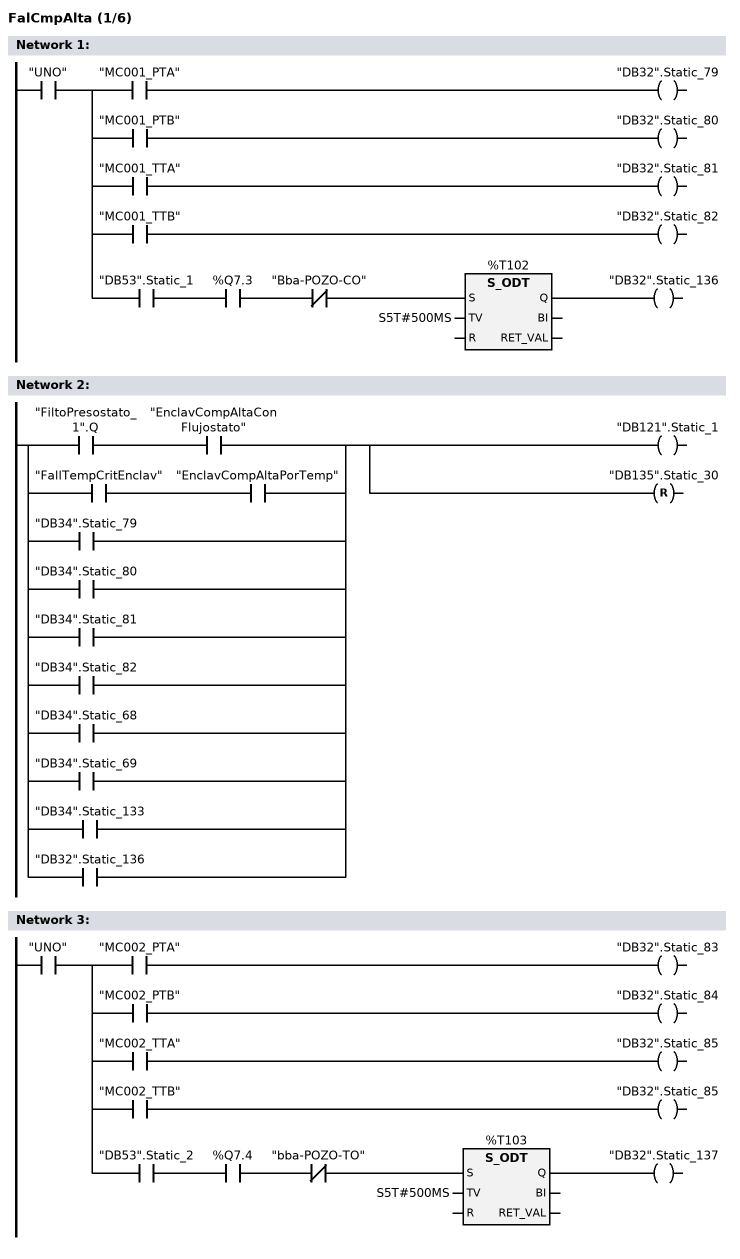
   RUNG wire#powerrail
      Contact( "UNO" )
      wire#w1
      Contact( "MC001_PTA" )
      Coil( "DB32".Static_79 )
   END_RUNG
   RUNG wire#w1
      Contact( "MC001_PTB" )
      Coil( "DB32".Static_80 )
   END_RUNG
   RUNG wire#w1
      Contact( "MC001_TTA" )
      Coil( "DB32".Static_81 )
   END_RUNG
   RUNG wire#w1
      Contact( "MC001_TTB" )
      Coil( "DB32".Static_82 )
   END_RUNG
   RUNG wire#w1
      Contact( "DB53".Static_1 )
      Contact( %Q7.3 )
      I_Contact( "Bba-POZO-CO" )
      S_ODT(T_NO := %T102, TV := S5T#500MS, R :=, BI =>, RET_VAL =>)
      Coil( "DB32".Static_136 )
   END_RUNG
   // the same network as SCL:
   "DB32".Static_79 := "UNO" AND "MC001_PTA";
   "DB32".Static_80 := "UNO" AND "MC001_PTB";
   "DB32".Static_81 := "UNO" AND "MC001_TTA";
   "DB32".Static_82 := "UNO" AND "MC001_TTB";
   #_s5time1 := S_ODT(T_NO := %T102,
                      TV := S5T#500MS,
                      S := "UNO" AND "DB53".Static_1 AND %Q7.3 AND NOT "Bba-POZO-CO",
                      Q => #_w1);
   "DB32".Static_136 := #_w1;
END_REGION

REGION Network 2
   "DB121".Static_1 := "DB34".Static_79 OR "DB34".Static_80 OR "DB34".Static_81 OR "DB34".Static_82 OR "DB34".Static_68 OR "DB34".Static_69 OR "DB34".Static_133 OR ("FiltoPresostato_1".Q AND "EnclavCompAltaConFlujostato") OR ("FallTempCritEnclav" AND "EnclavCompAltaPorTemp") OR "DB32".Static_136;
   IF "DB121".Static_1 THEN "DB135".Static_30 := FALSE; END_IF;
END_REGION

REGION Network 3
   RUNG wire#powerrail
      Contact( "UNO" )
      wire#w1
      Contact( "MC002_PTA" )
      Coil( "DB32".Static_83 )
   END_RUNG
   RUNG wire#w1
      Contact( "MC002_PTB" )
      Coil( "DB32".Static_84 )
   END_RUNG
   RUNG wire#w1
      Contact( "MC002_TTA" )
      Coil( "DB32".Static_85 )
   END_RUNG
   RUNG wire#w1
      Contact( "MC002_TTB" )
      Coil( "DB32".Static_85 )
   END_RUNG
   RUNG wire#w1
      Contact( "DB53".Static_2 )
      Contact( %Q7.4 )
      I_Contact( "bba-POZO-TO" )
      S_ODT(T_NO := %T103, TV := S5T#500MS, R :=, BI =>, RET_VAL =>)
      Coil( "DB32".Static_137 )
   END_RUNG
   // the same network as SCL:
   "DB32".Static_83 := "UNO" AND "MC002_PTA";
   "DB32".Static_84 := "UNO" AND "MC002_PTB";
   "DB32".Static_85 := "UNO" AND "MC002_TTA";
   "DB32".Static_85 := "UNO" AND "MC002_TTB";
   #_s5time1 := S_ODT(T_NO := %T103,
                      TV := S5T#500MS,
                      S := "UNO" AND "DB53".Static_2 AND %Q7.4 AND NOT "bba-POZO-TO",
                      Q => #_w1);
   "DB32".Static_137 := #_w1;
END_REGION

REGION Network 4
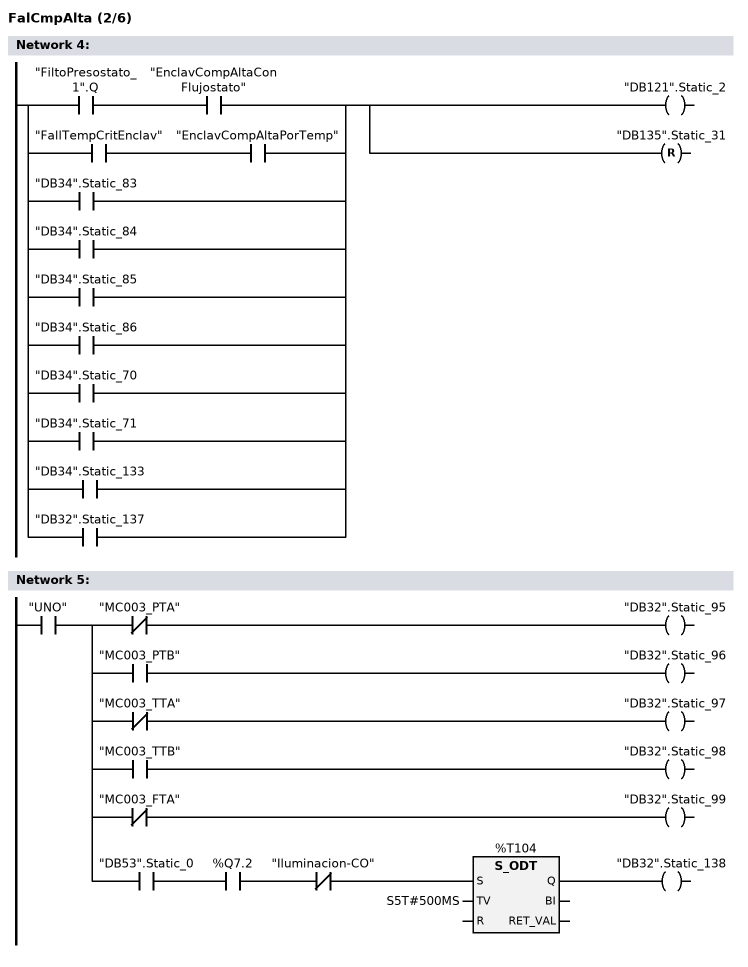
   "DB121".Static_2 := "DB34".Static_83 OR "DB34".Static_84 OR "DB34".Static_85 OR "DB34".Static_86 OR "DB34".Static_70 OR "DB34".Static_71 OR "DB34".Static_133 OR ("FiltoPresostato_1".Q AND "EnclavCompAltaConFlujostato") OR ("FallTempCritEnclav" AND "EnclavCompAltaPorTemp") OR "DB32".Static_137;
   IF "DB121".Static_2 THEN "DB135".Static_31 := FALSE; END_IF;
END_REGION

REGION Network 5
   RUNG wire#powerrail
      Contact( "UNO" )
      wire#w1
      I_Contact( "MC003_PTA" )
      Coil( "DB32".Static_95 )
   END_RUNG
   RUNG wire#w1
      Contact( "MC003_PTB" )
      Coil( "DB32".Static_96 )
   END_RUNG
   RUNG wire#w1
      I_Contact( "MC003_TTA" )
      Coil( "DB32".Static_97 )
   END_RUNG
   RUNG wire#w1
      Contact( "MC003_TTB" )
      Coil( "DB32".Static_98 )
   END_RUNG
   RUNG wire#w1
      I_Contact( "MC003_FTA" )
      Coil( "DB32".Static_99 )
   END_RUNG
   RUNG wire#w1
      Contact( "DB53".Static_0 )
      Contact( %Q7.2 )
      I_Contact( "Iluminacion-CO" )
      S_ODT(T_NO := %T104, TV := S5T#500MS, R :=, BI =>, RET_VAL =>)
      Coil( "DB32".Static_138 )
   END_RUNG
   // the same network as SCL:
   "DB32".Static_95 := "UNO" AND NOT "MC003_PTA";
   "DB32".Static_96 := "UNO" AND "MC003_PTB";
   "DB32".Static_97 := "UNO" AND NOT "MC003_TTA";
   "DB32".Static_98 := "UNO" AND "MC003_TTB";
   "DB32".Static_99 := "UNO" AND NOT "MC003_FTA";
   #_s5time1 := S_ODT(T_NO := %T104,
                      TV := S5T#500MS,
                      S := "UNO" AND "DB53".Static_0 AND %Q7.2 AND NOT "Iluminacion-CO",
                      Q => #_w1);
   "DB32".Static_138 := #_w1;
END_REGION

REGION Network 6
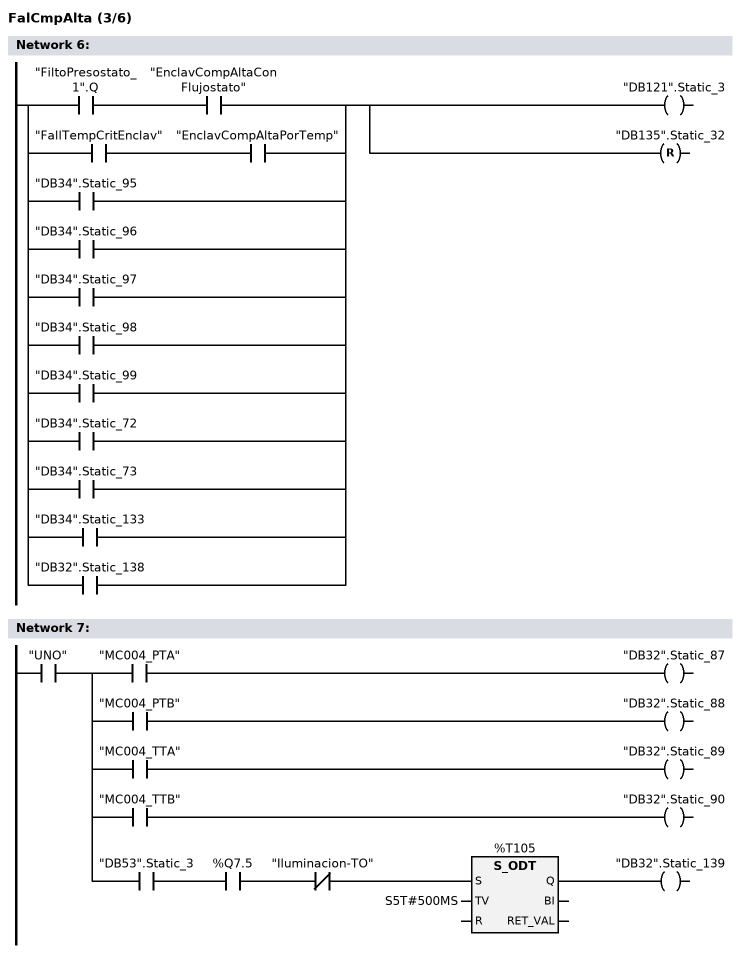
   "DB121".Static_3 := "DB34".Static_95 OR "DB34".Static_96 OR "DB34".Static_97 OR "DB34".Static_98 OR "DB34".Static_99 OR "DB34".Static_72 OR "DB34".Static_73 OR "DB34".Static_133 OR ("FiltoPresostato_1".Q AND "EnclavCompAltaConFlujostato") OR ("FallTempCritEnclav" AND "EnclavCompAltaPorTemp") OR "DB32".Static_138;
   IF "DB121".Static_3 THEN "DB135".Static_32 := FALSE; END_IF;
END_REGION

REGION Network 7
   RUNG wire#powerrail
      Contact( "UNO" )
      wire#w1
      Contact( "MC004_PTA" )
      Coil( "DB32".Static_87 )
   END_RUNG
   RUNG wire#w1
      Contact( "MC004_PTB" )
      Coil( "DB32".Static_88 )
   END_RUNG
   RUNG wire#w1
      Contact( "MC004_TTA" )
      Coil( "DB32".Static_89 )
   END_RUNG
   RUNG wire#w1
      Contact( "MC004_TTB" )
      Coil( "DB32".Static_90 )
   END_RUNG
   RUNG wire#w1
      Contact( "DB53".Static_3 )
      Contact( %Q7.5 )
      I_Contact( "Iluminacion-TO" )
      S_ODT(T_NO := %T105, TV := S5T#500MS, R :=, BI =>, RET_VAL =>)
      Coil( "DB32".Static_139 )
   END_RUNG
   // the same network as SCL:
   "DB32".Static_87 := "UNO" AND "MC004_PTA";
   "DB32".Static_88 := "UNO" AND "MC004_PTB";
   "DB32".Static_89 := "UNO" AND "MC004_TTA";
   "DB32".Static_90 := "UNO" AND "MC004_TTB";
   #_s5time1 := S_ODT(T_NO := %T105,
                      TV := S5T#500MS,
                      S := "UNO" AND "DB53".Static_3 AND %Q7.5 AND NOT "Iluminacion-TO",
                      Q => #_w1);
   "DB32".Static_139 := #_w1;
END_REGION

REGION Network 8
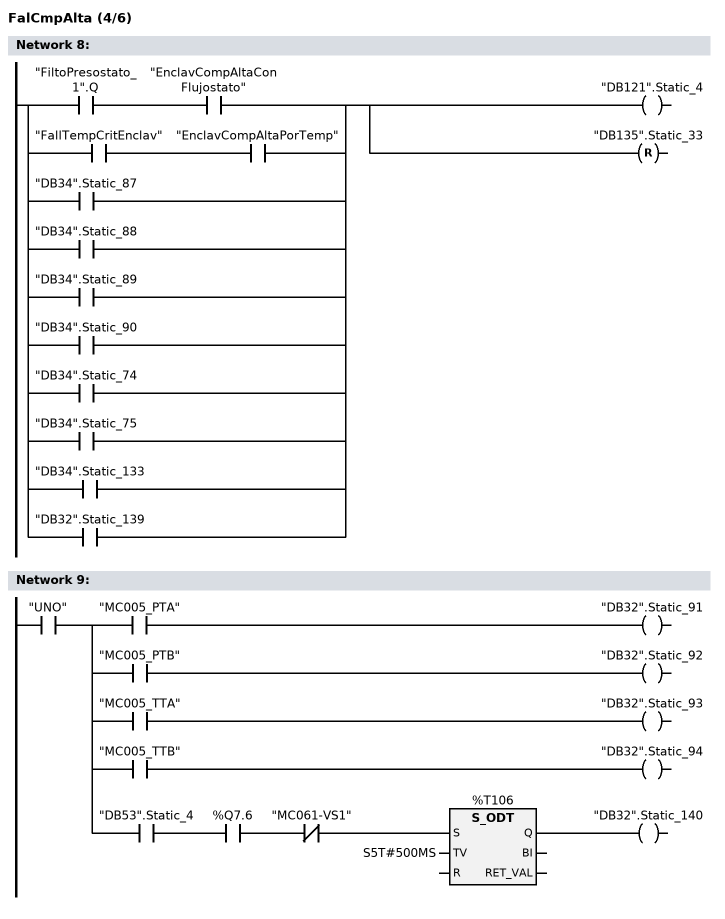
   "DB121".Static_4 := "DB34".Static_87 OR "DB34".Static_88 OR "DB34".Static_89 OR "DB34".Static_90 OR "DB34".Static_74 OR "DB34".Static_75 OR "DB34".Static_133 OR ("FiltoPresostato_1".Q AND "EnclavCompAltaConFlujostato") OR ("FallTempCritEnclav" AND "EnclavCompAltaPorTemp") OR "DB32".Static_139;
   IF "DB121".Static_4 THEN "DB135".Static_33 := FALSE; END_IF;
END_REGION

REGION Network 9
   RUNG wire#powerrail
      Contact( "UNO" )
      wire#w1
      Contact( "MC005_PTA" )
      Coil( "DB32".Static_91 )
   END_RUNG
   RUNG wire#w1
      Contact( "MC005_PTB" )
      Coil( "DB32".Static_92 )
   END_RUNG
   RUNG wire#w1
      Contact( "MC005_TTA" )
      Coil( "DB32".Static_93 )
   END_RUNG
   RUNG wire#w1
      Contact( "MC005_TTB" )
      Coil( "DB32".Static_94 )
   END_RUNG
   RUNG wire#w1
      Contact( "DB53".Static_4 )
      Contact( %Q7.6 )
      I_Contact( "MC061-VS1" )
      S_ODT(T_NO := %T106, TV := S5T#500MS, R :=, BI =>, RET_VAL =>)
      Coil( "DB32".Static_140 )
   END_RUNG
   // the same network as SCL:
   "DB32".Static_91 := "UNO" AND "MC005_PTA";
   "DB32".Static_92 := "UNO" AND "MC005_PTB";
   "DB32".Static_93 := "UNO" AND "MC005_TTA";
   "DB32".Static_94 := "UNO" AND "MC005_TTB";
   #_s5time1 := S_ODT(T_NO := %T106,
                      TV := S5T#500MS,
                      S := "UNO" AND "DB53".Static_4 AND %Q7.6 AND NOT "MC061-VS1",
                      Q => #_w1);
   "DB32".Static_140 := #_w1;
END_REGION

REGION Network 10
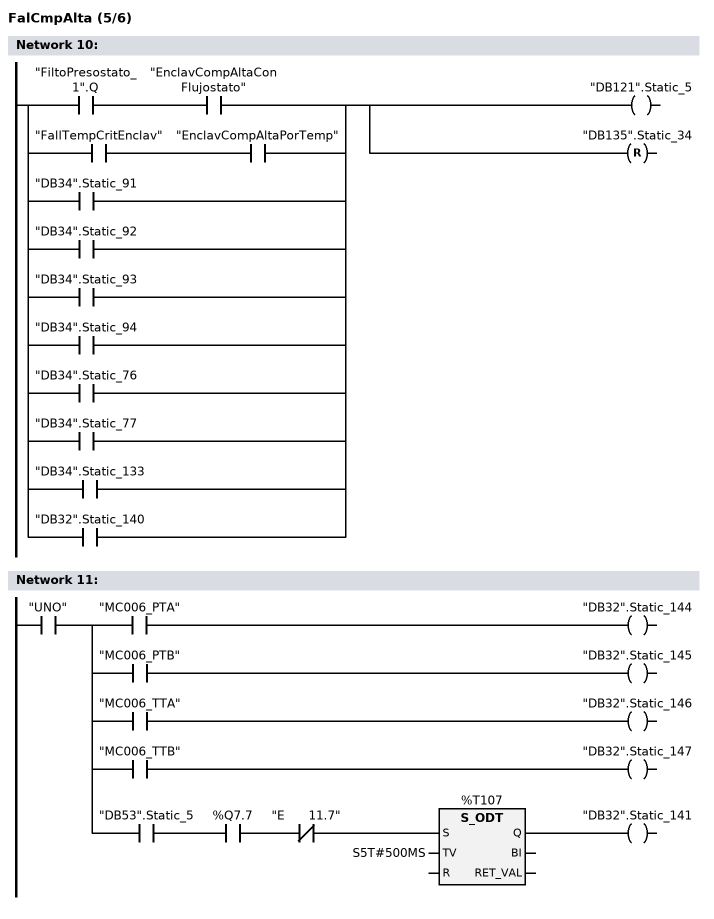
   "DB121".Static_5 := "DB34".Static_91 OR "DB34".Static_92 OR "DB34".Static_93 OR "DB34".Static_94 OR "DB34".Static_76 OR "DB34".Static_77 OR "DB34".Static_133 OR ("FiltoPresostato_1".Q AND "EnclavCompAltaConFlujostato") OR ("FallTempCritEnclav" AND "EnclavCompAltaPorTemp") OR "DB32".Static_140;
   IF "DB121".Static_5 THEN "DB135".Static_34 := FALSE; END_IF;
END_REGION

REGION Network 11
   RUNG wire#powerrail
      Contact( "UNO" )
      wire#w1
      Contact( "MC006_PTA" )
      Coil( "DB32".Static_144 )
   END_RUNG
   RUNG wire#w1
      Contact( "MC006_PTB" )
      Coil( "DB32".Static_145 )
   END_RUNG
   RUNG wire#w1
      Contact( "MC006_TTA" )
      Coil( "DB32".Static_146 )
   END_RUNG
   RUNG wire#w1
      Contact( "MC006_TTB" )
      Coil( "DB32".Static_147 )
   END_RUNG
   RUNG wire#w1
      Contact( "DB53".Static_5 )
      Contact( %Q7.7 )
      I_Contact( "E      11.7" )
      S_ODT(T_NO := %T107, TV := S5T#500MS, R :=, BI =>, RET_VAL =>)
      Coil( "DB32".Static_141 )
   END_RUNG
   // the same network as SCL:
   "DB32".Static_144 := "UNO" AND "MC006_PTA";
   "DB32".Static_145 := "UNO" AND "MC006_PTB";
   "DB32".Static_146 := "UNO" AND "MC006_TTA";
   "DB32".Static_147 := "UNO" AND "MC006_TTB";
   #_s5time1 := S_ODT(T_NO := %T107,
                      TV := S5T#500MS,
                      S := "UNO" AND "DB53".Static_5 AND %Q7.7 AND NOT "E      11.7",
                      Q => #_w1);
   "DB32".Static_141 := #_w1;
END_REGION

REGION Network 12
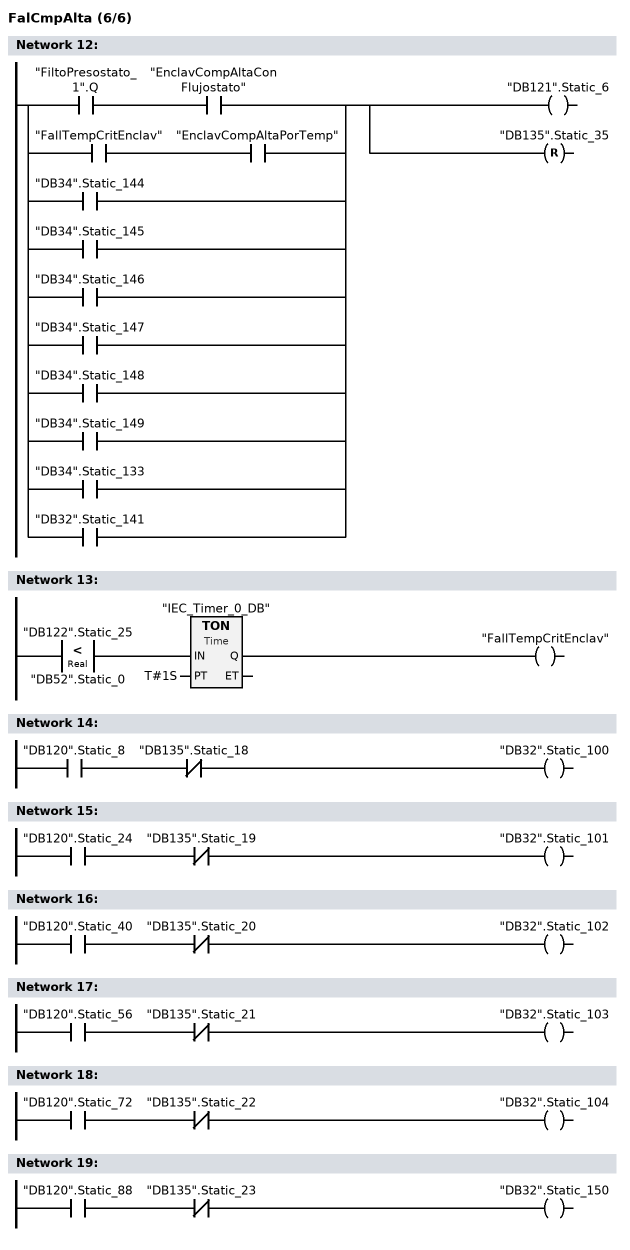
   "DB121".Static_6 := "DB34".Static_144 OR "DB34".Static_145 OR "DB34".Static_146 OR "DB34".Static_147 OR "DB34".Static_148 OR "DB34".Static_149 OR "DB34".Static_133 OR ("FiltoPresostato_1".Q AND "EnclavCompAltaConFlujostato") OR ("FallTempCritEnclav" AND "EnclavCompAltaPorTemp") OR "DB32".Static_141;
   IF "DB121".Static_6 THEN "DB135".Static_35 := FALSE; END_IF;
END_REGION

REGION Network 13
   "IEC_Timer_0_DB".TON(in := "DB122".Static_25 < "DB52".Static_0, pt := T#1S);
   "FallTempCritEnclav" := "IEC_Timer_0_DB".q;
END_REGION

REGION Network 14
   RUNG wire#powerrail
      Contact( "DB120".Static_8 )
      I_Contact( "DB135".Static_18 )
      Coil( "DB32".Static_100 )
   END_RUNG
   // the same network as SCL:
   "DB32".Static_100 := "DB120".Static_8 AND NOT "DB135".Static_18;
END_REGION

REGION Network 15
   RUNG wire#powerrail
      Contact( "DB120".Static_24 )
      I_Contact( "DB135".Static_19 )
      Coil( "DB32".Static_101 )
   END_RUNG
   // the same network as SCL:
   "DB32".Static_101 := "DB120".Static_24 AND NOT "DB135".Static_19;
END_REGION

REGION Network 16
   RUNG wire#powerrail
      Contact( "DB120".Static_40 )
      I_Contact( "DB135".Static_20 )
      Coil( "DB32".Static_102 )
   END_RUNG
   // the same network as SCL:
   "DB32".Static_102 := "DB120".Static_40 AND NOT "DB135".Static_20;
END_REGION

REGION Network 17
   RUNG wire#powerrail
      Contact( "DB120".Static_56 )
      I_Contact( "DB135".Static_21 )
      Coil( "DB32".Static_103 )
   END_RUNG
   // the same network as SCL:
   "DB32".Static_103 := "DB120".Static_56 AND NOT "DB135".Static_21;
END_REGION

REGION Network 18
   RUNG wire#powerrail
      Contact( "DB120".Static_72 )
      I_Contact( "DB135".Static_22 )
      Coil( "DB32".Static_104 )
   END_RUNG
   // the same network as SCL:
   "DB32".Static_104 := "DB120".Static_72 AND NOT "DB135".Static_22;
END_REGION

REGION Network 19
   RUNG wire#powerrail
      Contact( "DB120".Static_88 )
      I_Contact( "DB135".Static_23 )
      Coil( "DB32".Static_150 )
   END_RUNG
   // the same network as SCL:
   "DB32".Static_150 := "DB120".Static_88 AND NOT "DB135".Static_23;
END_REGION
END_FUNCTION

// folder: Auxiliares

FUNCTION "AjusteEntrada-SalidaMTA" : Void   // FC6, LAD
{ S7_Optimized_Access := 'FALSE' }
VERSION : 0.1
BEGIN

REGION Network 1
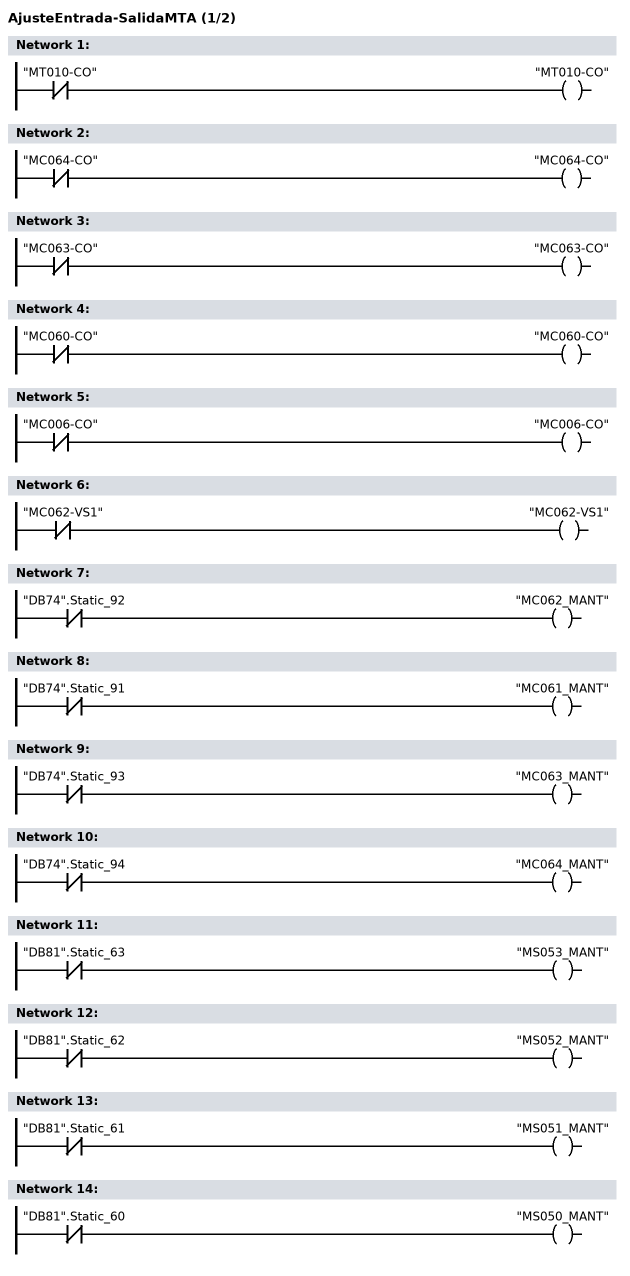
   RUNG wire#powerrail
      I_Contact( "MT010-CO" )
      Coil( "MT010-CO" )
   END_RUNG
   // the same network as SCL:
   "MT010-CO" := NOT "MT010-CO";
END_REGION

REGION Network 2
   RUNG wire#powerrail
      I_Contact( "MC064-CO" )
      Coil( "MC064-CO" )
   END_RUNG
   // the same network as SCL:
   "MC064-CO" := NOT "MC064-CO";
END_REGION

REGION Network 3
   RUNG wire#powerrail
      I_Contact( "MC063-CO" )
      Coil( "MC063-CO" )
   END_RUNG
   // the same network as SCL:
   "MC063-CO" := NOT "MC063-CO";
END_REGION

REGION Network 4
   RUNG wire#powerrail
      I_Contact( "MC060-CO" )
      Coil( "MC060-CO" )
   END_RUNG
   // the same network as SCL:
   "MC060-CO" := NOT "MC060-CO";
END_REGION

REGION Network 5
   RUNG wire#powerrail
      I_Contact( "MC006-CO" )
      Coil( "MC006-CO" )
   END_RUNG
   // the same network as SCL:
   "MC006-CO" := NOT "MC006-CO";
END_REGION

REGION Network 6
   RUNG wire#powerrail
      I_Contact( "MC062-VS1" )
      Coil( "MC062-VS1" )
   END_RUNG
   // the same network as SCL:
   "MC062-VS1" := NOT "MC062-VS1";
END_REGION

REGION Network 7
   RUNG wire#powerrail
      I_Contact( "DB74".Static_92 )
      Coil( "MC062_MANT" )
   END_RUNG
   // the same network as SCL:
   "MC062_MANT" := NOT "DB74".Static_92;
END_REGION

REGION Network 8
   RUNG wire#powerrail
      I_Contact( "DB74".Static_91 )
      Coil( "MC061_MANT" )
   END_RUNG
   // the same network as SCL:
   "MC061_MANT" := NOT "DB74".Static_91;
END_REGION

REGION Network 9
   RUNG wire#powerrail
      I_Contact( "DB74".Static_93 )
      Coil( "MC063_MANT" )
   END_RUNG
   // the same network as SCL:
   "MC063_MANT" := NOT "DB74".Static_93;
END_REGION

REGION Network 10
   RUNG wire#powerrail
      I_Contact( "DB74".Static_94 )
      Coil( "MC064_MANT" )
   END_RUNG
   // the same network as SCL:
   "MC064_MANT" := NOT "DB74".Static_94;
END_REGION

REGION Network 11
   RUNG wire#powerrail
      I_Contact( "DB81".Static_63 )
      Coil( "MS053_MANT" )
   END_RUNG
   // the same network as SCL:
   "MS053_MANT" := NOT "DB81".Static_63;
END_REGION

REGION Network 12
   RUNG wire#powerrail
      I_Contact( "DB81".Static_62 )
      Coil( "MS052_MANT" )
   END_RUNG
   // the same network as SCL:
   "MS052_MANT" := NOT "DB81".Static_62;
END_REGION

REGION Network 13
   RUNG wire#powerrail
      I_Contact( "DB81".Static_61 )
      Coil( "MS051_MANT" )
   END_RUNG
   // the same network as SCL:
   "MS051_MANT" := NOT "DB81".Static_61;
END_REGION

REGION Network 14
   RUNG wire#powerrail
      I_Contact( "DB81".Static_60 )
      Coil( "MS050_MANT" )
   END_RUNG
   // the same network as SCL:
   "MS050_MANT" := NOT "DB81".Static_60;
END_REGION

REGION Network 15
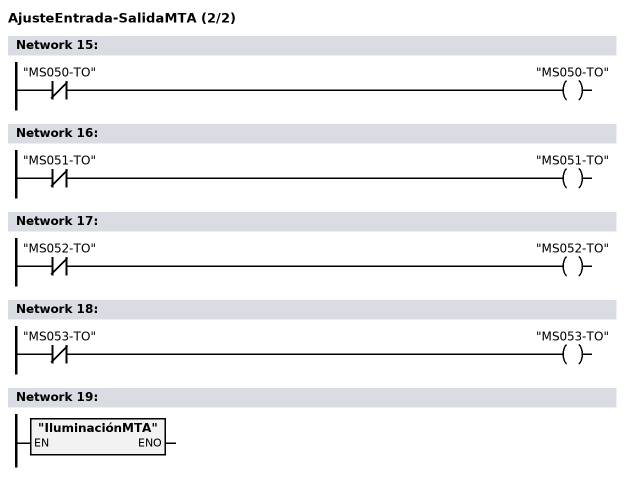
   RUNG wire#powerrail
      I_Contact( "MS050-TO" )
      Coil( "MS050-TO" )
   END_RUNG
   // the same network as SCL:
   "MS050-TO" := NOT "MS050-TO";
END_REGION

REGION Network 16
   RUNG wire#powerrail
      I_Contact( "MS051-TO" )
      Coil( "MS051-TO" )
   END_RUNG
   // the same network as SCL:
   "MS051-TO" := NOT "MS051-TO";
END_REGION

REGION Network 17
   RUNG wire#powerrail
      I_Contact( "MS052-TO" )
      Coil( "MS052-TO" )
   END_RUNG
   // the same network as SCL:
   "MS052-TO" := NOT "MS052-TO";
END_REGION

REGION Network 18
   RUNG wire#powerrail
      I_Contact( "MS053-TO" )
      Coil( "MS053-TO" )
   END_RUNG
   // the same network as SCL:
   "MS053-TO" := NOT "MS053-TO";
END_REGION

REGION Network 19
   RUNG wire#powerrail
      "IluminaciónMTA"()
   END_RUNG
   // the same network as SCL:
   "IluminaciónMTA"();
END_REGION
END_FUNCTION

FUNCTION "And-Byte MTA" : Void   // FC22, LAD
{ S7_Optimized_Access := 'FALSE' }
VERSION : 0.1
BEGIN

REGION Network 1
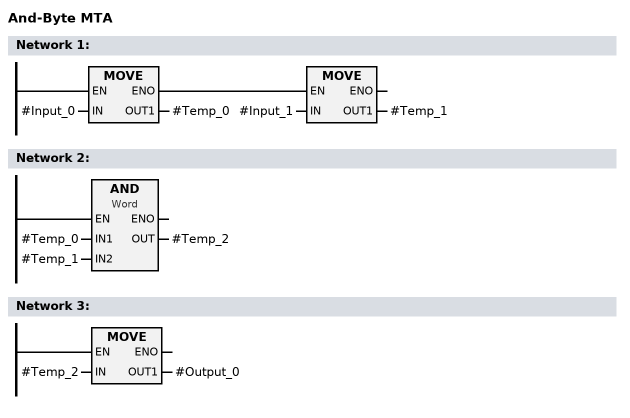
   RUNG wire#powerrail
      { S7_GenerateENO := "TRUE" } Move(in := #Input_0, out1 => #Temp_0)
      { S7_GenerateENO := "TRUE" } Move(in := #Input_1, out1 => #Temp_1)
   END_RUNG
   // the same network as SCL:
   // ENO of a box is taken as its EN; it also drops when the box reports an error
   #Temp_0 := #Input_0;
   #Temp_1 := #Input_1;
END_REGION

REGION Network 2
   RUNG wire#powerrail
      { S7_Templates := "SrcType := Word"; S7_GenerateENO := "TRUE" } And(in1 := #Temp_0, in2 := #Temp_1, out => #Temp_2)
   END_RUNG
   // the same network as SCL:
   #Temp_2 := #Temp_0 AND #Temp_1;
END_REGION

REGION Network 3
   RUNG wire#powerrail
      { S7_GenerateENO := "TRUE" } Move(in := #Temp_2, out1 => #Output_0)
   END_RUNG
   // the same network as SCL:
   #Output_0 := #Temp_2;
END_REGION
END_FUNCTION

FUNCTION "Inicialización" : Void   // FC46, LAD
{ S7_Optimized_Access := 'FALSE' }
VERSION : 0.1
BEGIN

REGION Network 1
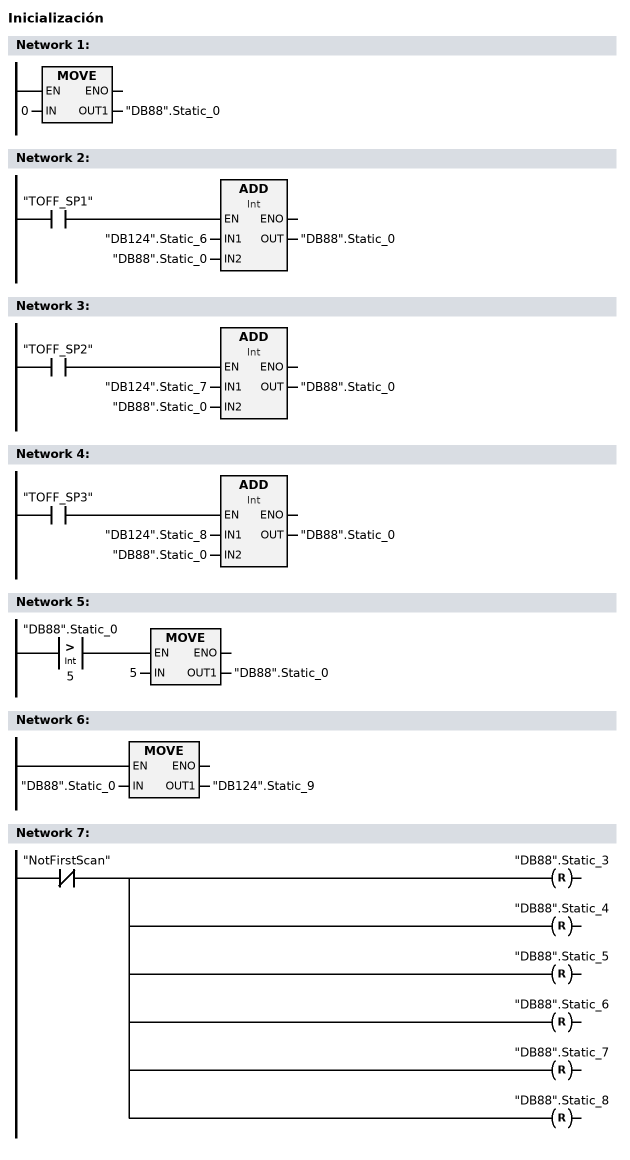
   RUNG wire#powerrail
      { S7_GenerateENO := "TRUE" } Move(in := 0, out1 => "DB88".Static_0)
   END_RUNG
   // the same network as SCL:
   "DB88".Static_0 := 0;
END_REGION

REGION Network 2
   RUNG wire#powerrail
      Contact( "TOFF_SP1" )
      { S7_Templates := "SrcType := Int"; S7_GenerateENO := "TRUE" } Add(in1 := "DB124".Static_6, in2 := "DB88".Static_0, out => "DB88".Static_0)
   END_RUNG
   // the same network as SCL:
   IF "TOFF_SP1" THEN "DB88".Static_0 := "DB124".Static_6 + "DB88".Static_0; END_IF;
END_REGION

REGION Network 3
   RUNG wire#powerrail
      Contact( "TOFF_SP2" )
      { S7_Templates := "SrcType := Int"; S7_GenerateENO := "TRUE" } Add(in1 := "DB124".Static_7, in2 := "DB88".Static_0, out => "DB88".Static_0)
   END_RUNG
   // the same network as SCL:
   IF "TOFF_SP2" THEN "DB88".Static_0 := "DB124".Static_7 + "DB88".Static_0; END_IF;
END_REGION

REGION Network 4
   RUNG wire#powerrail
      Contact( "TOFF_SP3" )
      { S7_Templates := "SrcType := Int"; S7_GenerateENO := "TRUE" } Add(in1 := "DB124".Static_8, in2 := "DB88".Static_0, out => "DB88".Static_0)
   END_RUNG
   // the same network as SCL:
   IF "TOFF_SP3" THEN "DB88".Static_0 := "DB124".Static_8 + "DB88".Static_0; END_IF;
END_REGION

REGION Network 5
   RUNG wire#powerrail
      { S7_Templates := "SrcType := Int" } GT_Contact(in1 := "DB88".Static_0, in2 := 5)
      { S7_GenerateENO := "TRUE" } Move(in := 5, out1 => "DB88".Static_0)
   END_RUNG
   // the same network as SCL:
   IF "DB88".Static_0 > 5 THEN "DB88".Static_0 := 5; END_IF;
END_REGION

REGION Network 6
   RUNG wire#powerrail
      { S7_GenerateENO := "TRUE" } Move(in := "DB88".Static_0, out1 => "DB124".Static_9)
   END_RUNG
   // the same network as SCL:
   "DB124".Static_9 := "DB88".Static_0;
END_REGION

REGION Network 7
   RUNG wire#powerrail
      I_Contact( "NotFirstScan" )
      wire#w1
      R_Coil( "DB88".Static_3 )
   END_RUNG
   RUNG wire#w1
      R_Coil( "DB88".Static_4 )
   END_RUNG
   RUNG wire#w1
      R_Coil( "DB88".Static_5 )
   END_RUNG
   RUNG wire#w1
      R_Coil( "DB88".Static_6 )
   END_RUNG
   RUNG wire#w1
      R_Coil( "DB88".Static_7 )
   END_RUNG
   RUNG wire#w1
      R_Coil( "DB88".Static_8 )
   END_RUNG
   // the same network as SCL:
   IF NOT "NotFirstScan" THEN
       "DB88".Static_3 := FALSE;
       "DB88".Static_4 := FALSE;
       "DB88".Static_5 := FALSE;
       "DB88".Static_6 := FALSE;
       "DB88".Static_7 := FALSE;
       "DB88".Static_8 := FALSE;
   END_IF;
END_REGION
END_FUNCTION

// folder: Bloques Estandar

FUNCTION_BLOCK "ControladorMotoresMTA"   // FB2, LAD
{ S7_Optimized_Access := 'FALSE' }
VERSION : 0.1
BEGIN

REGION Network 2
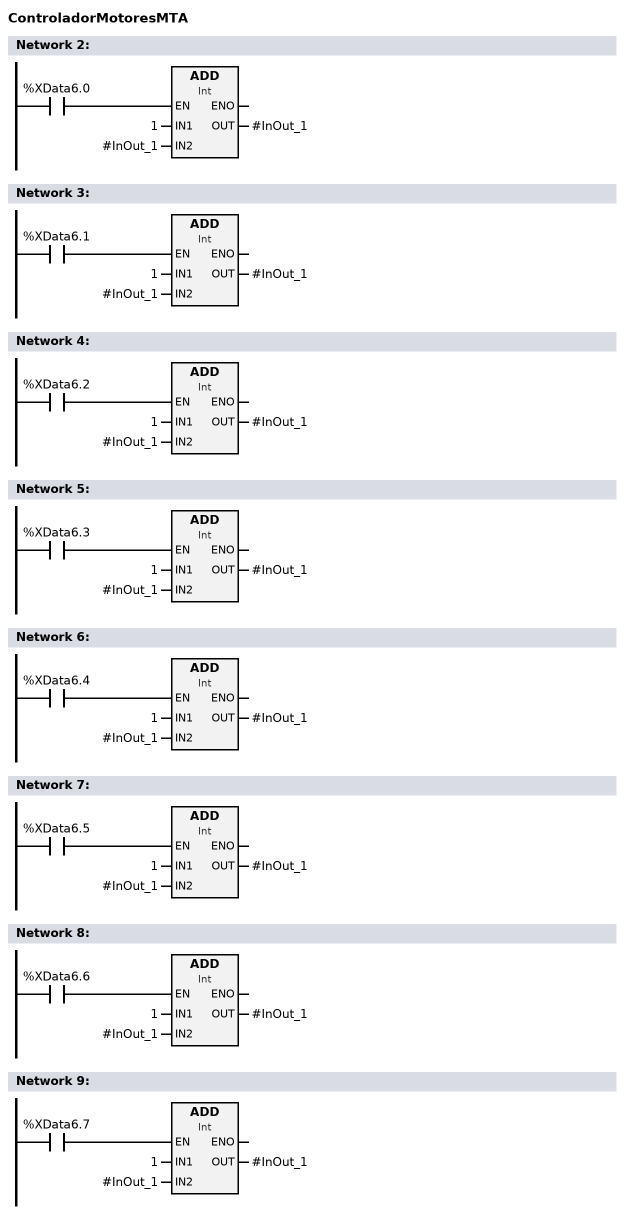
   RUNG wire#powerrail
      Contact( %XData6.0 )
      { S7_Templates := "SrcType := Int"; S7_GenerateENO := "TRUE" } Add(in1 := 1, in2 := #InOut_1, out => #InOut_1)
   END_RUNG
   // the same network as SCL:
   IF %XData6.0 THEN #InOut_1 := 1 + #InOut_1; END_IF;
END_REGION

REGION Network 3
   RUNG wire#powerrail
      Contact( %XData6.1 )
      { S7_Templates := "SrcType := Int"; S7_GenerateENO := "TRUE" } Add(in1 := 1, in2 := #InOut_1, out => #InOut_1)
   END_RUNG
   // the same network as SCL:
   IF %XData6.1 THEN #InOut_1 := 1 + #InOut_1; END_IF;
END_REGION

REGION Network 4
   RUNG wire#powerrail
      Contact( %XData6.2 )
      { S7_Templates := "SrcType := Int"; S7_GenerateENO := "TRUE" } Add(in1 := 1, in2 := #InOut_1, out => #InOut_1)
   END_RUNG
   // the same network as SCL:
   IF %XData6.2 THEN #InOut_1 := 1 + #InOut_1; END_IF;
END_REGION

REGION Network 5
   RUNG wire#powerrail
      Contact( %XData6.3 )
      { S7_Templates := "SrcType := Int"; S7_GenerateENO := "TRUE" } Add(in1 := 1, in2 := #InOut_1, out => #InOut_1)
   END_RUNG
   // the same network as SCL:
   IF %XData6.3 THEN #InOut_1 := 1 + #InOut_1; END_IF;
END_REGION

REGION Network 6
   RUNG wire#powerrail
      Contact( %XData6.4 )
      { S7_Templates := "SrcType := Int"; S7_GenerateENO := "TRUE" } Add(in1 := 1, in2 := #InOut_1, out => #InOut_1)
   END_RUNG
   // the same network as SCL:
   IF %XData6.4 THEN #InOut_1 := 1 + #InOut_1; END_IF;
END_REGION

REGION Network 7
   RUNG wire#powerrail
      Contact( %XData6.5 )
      { S7_Templates := "SrcType := Int"; S7_GenerateENO := "TRUE" } Add(in1 := 1, in2 := #InOut_1, out => #InOut_1)
   END_RUNG
   // the same network as SCL:
   IF %XData6.5 THEN #InOut_1 := 1 + #InOut_1; END_IF;
END_REGION
